   "DB_Inspect_Pistoane_PompaB" : Int = PLC DB_Inspect_Pistoane.Piston_A AT %DB34.DBW28, 1 s
   "DB_Inspect_Pistoane_PompaC" : Int = PLC DB_Inspect_Pistoane.Piston_B AT %DB34.DBW30, 1 s
   "DB_Inspect_Pistoane_CutP1" : Bool = PLC DB_Inspect_Pistoane.Piston_C AT %DB34.DBX32.5, 1 s
   "DB_Inspect_Pistoane_StatusPump1" : Int = PLC DB_Inspect_Pistoane.Presiune_1 AT %DB34.DBW34, 1 s
   "DB_Vizibilitati_Platforme/Colete_Platforma_Rebut" : Bool = PLC DB_Inspect_Pistoane.Presiune_2 AT %DB1.DBX1.0, 100 ms
   "DB_Vizibilitati_Platforme/Colete_Colet_Rebut" : Bool = PLC DB_Inspect_Pistoane.Presiune_A AT %DB1.DBX0.7, 100 ms
   "DB_Tip_Cutie_BoxStatus" : Bool = PLC DB_Inspect_Pistoane.Presiune_B AT %DB37.DBX6.3, 100 ms
   "DB_ControlEnable_ControlEnable_Btn_A" : Bool = PLC DB_Inspect_Pistoane.Presiune_C AT %DB45.DBX0.0, 1 s
   "DB_ControlEnable_ControlEnable_Btn_B" : Bool = PLC DB_Inspect_Pistoane.Presiune_Upper_2 AT %DB45.DBX0.1, 1 s
   "DB_ControlEnable_ControlEnable_Btn_C" : Bool = PLC DB_Inspect_Pistoane.Presiune_Upper_1 AT %DB45.DBX0.2, 1 s
   "DB_ControlEnable_ControlEnable_Btn_Load" : Bool = PLC DB_Inspect_Pistoane.Presiune_Lower_1 AT %DB45.DBX0.3, 1 s
   "DB_ControlEnable_ControlEnable_Btn_ACKLoad" : Bool = PLC DB_Inspect_Pistoane.Presiune_Lower_2 AT %DB45.DBX0.4, 1 s
   "DB_ControlEnable_ControlEnable_Btn_PlaceBox" : Bool = PLC DB_Status_Motoare.Motor_1 AT %DB45.DBX0.6, 1 s
   "DB_general_Piston_Scrap" : Int = PLC DB_HMI.Viz_Platforma_Libera AT %DB2.DBW36, 100 ms
   "DB_Tranzitii_Viz_CutieScrapP3" : Bool = PLC DB_general.Piston_Incarcare AT %DB47.DBX8.0, 100 ms
   "DB_Banda3_AckScrap" : Bool = PLC DB_Banda3.AckScrap AT %DB49.DBX2.1, 100 ms
   "DB_Banda3_Poz_Banda3" : Int = PLC DB_Banda3.Poz_Banda3 AT %DB49.DBW0, 100 ms
   "DB_Banda3_Viz_CutieBanda3" : Bool = PLC DB_Banda3.Viz_CutieBanda3 AT %DB49.DBX2.0, 100 ms
   "DB_HMI_Eng/Ger" : Bool = PLC DB_HMI.Eng AT %DB19.DBX124.0, 1 s
   "DB_HMI_Ger" : Bool = PLC DB_HMI.Ger AT %DB19.DBX138.0, 1 s
   "DB_RemoteAcces_ControlEnable_Stop" : Bool = PLC DB_RemoteAcces.ControlEnable_Stop AT %DB6.DBX0.6, 1 s
   "DB_RemoteAcces_ControlEnable_Start" : Bool = PLC DB_RemoteAcces.ControlEnable_Start AT %DB6.DBX0.7, 1 s
   "DB_RemoteAcces_ControlEnable_Man/Auto" : Bool = PLC DB_RemoteAcces.ControlEnable_Man/Auto AT %DB6.DBX1.0, 1 s
   "DB_ControlEnable_ControlEnable_StartSim" : Bool = PLC DB_ControlEnable.ControlEnable_StartSim AT %DB45.DBX0.5, 1 s
   "DB_SIM_Ack_Load_Pressed" : Bool = PLC DB_SIM.Ack_Load_Pressed AT %DB40.DBX0.3, 1 s
   "DB_ControlEnable_StatusLoadBtn" : Int = PLC DB_ControlEnable.StatusLoadBtn AT %DB45.DBW2, 1 s

HMI tags "Vizibilitate_Log"
   "Viz_Pachet_1" : Bool, internal
   "Viz_Pachet_2" : Bool, internal
   "Viz_Pachet_3" : Bool, internal
   "Viz_Pachet_4" : Bool, internal
   "Viz_Pachet_5" : Bool, internal
   "Viz_Pachet_6" : Bool, internal
   "Viz_Pachet_7" : Bool, internal
   "Viz_Pachet_8" : Bool, internal
   "Viz_Pachet_9" : Bool, internal
   "Viz_Pachet_10" : Bool, internal
   "QR_En" : Bool, internal

HMI tags "DB_HMI_tags"
   "DB_HMI_A_Pressed" : Bool = PLC DB_HMI.A_Pressed AT %DB19.DBX6.0, 100 ms
   "DB_HMI_Ack_Load" : Bool = PLC DB_HMI.Ack_Load AT %DB19.DBX14.3, 100 ms
   "DB_HMI_Add_Ulei" : Bool = PLC DB_HMI.Add_Ulei AT %DB19.DBX42.0, 100 ms
   "DB_HMI_B_Pressed" : Bool = PLC DB_HMI.B_Pressed AT %DB19.DBX6.1, 100 ms
   "DB_HMI_C_Pressed" : Bool = PLC DB_HMI.C_Pressed AT %DB19.DBX6.2, 100 ms
   "DB_HMI_Cutie_Automata" : Bool = PLC DB_HMI.Cutie_Automata AT %DB19.DBX6.3, 100 ms
   "DB_HMI_Cutie_Manuala" : Bool = PLC DB_HMI.Cutie_Manuala AT %DB19.DBX6.4, 100 ms
   "DB_HMI_Greutate" : Real = PLC DB_HMI.Greutate AT %DB19.DBD54, 100 ms
   "DB_HMI_LOAD" : Int = PLC DB_HMI.LOAD AT %DB19.DBW12, 100 ms
   "DB_HMI_LOAD_A" : Bool = PLC DB_HMI.LOAD_A AT %DB19.DBX28.0, 100 ms
   "DB_HMI_LOAD_B" : Bool = PLC DB_HMI.LOAD_B AT %DB19.DBX28.1, 100 ms
   "DB_HMI_LOAD_C" : Bool = PLC DB_HMI.LOAD_C AT %DB19.DBX28.2, 100 ms
   "DB_HMI_Load_RDY" : Bool = PLC DB_HMI.Load_RDY AT %DB19.DBX20.0, 100 ms
   "DB_HMI_Piston_1_Status" : Int = PLC DB_HMI.Piston_1_Status AT %DB19.DBW16, 100 ms
   "DB_HMI_Piston_2_Status" : Int = PLC DB_HMI.Piston_2_Status AT %DB19.DBW18, 100 ms
   "DB_HMI_Racire_Ulei" : Bool = PLC DB_HMI.Racire_Ulei AT %DB19.DBX42.3, 100 ms
   "DB_HMI_Sageata_Deplasare_Banda_Bile" : Bool = PLC DB_HMI.Sageata_Deplasare_Banda_Bile AT %DB19.DBX32.0, 100 ms
   "DB_HMI_Set_T0" : Bool = PLC DB_HMI.Set_T0 AT %DB19.DBX42.6, 100 ms
   "DB_HMI_Set_T50" : Bool = PLC DB_HMI.Set_T50 AT %DB19.DBX42.7, 100 ms
   "DB_HMI_START_SIM" : Bool = PLC DB_HMI.START_SIM AT %DB19.DBX43.0, 100 ms
   "DB_HMI_Start_System" : Bool = PLC DB_HMI.Start_System AT %DB19.DBX42.2, 100 ms
   "DB_HMI_Status_Banda_Bile" : Int = PLC DB_HMI.Status_Banda_Bile AT %DB19.DBW30, 100 ms
   "DB_HMI_Status_Incalzire/Racire_Ulei" : Int = PLC DB_HMI.Status_Incalzire/Racire_Ulei AT %DB19.DBW44, 100 ms
   "DB_HMI_Status_Piston_A" : Int = PLC DB_HMI.Status_Piston_A AT %DB19.DBW22, 100 ms
   "DB_HMI_Status_Piston_B" : Int = PLC DB_HMI.Status_Piston_B AT %DB19.DBW24, 100 ms
   "DB_HMI_Status_Piston_C" : Int = PLC DB_HMI.Status_Piston_C AT %DB19.DBW26, 100 ms
   "DB_HMI_Sub_Ulei" : Bool = PLC DB_HMI.Sub_Ulei AT %DB19.DBX42.1, 100 ms
   "DB_HMI_Temp_Ulei" : Int = PLC DB_HMI.Temp_Ulei AT %DB19.DBW34, 100 ms
   "DB_HMI_TEST_LOAD" : Bool = PLC DB_HMI.BTN_LOAD AT %DB19.DBX43.1, 100 ms
   "DB_HMI_Tip_Cutie" : Int = PLC DB_HMI.Tip_Cutie_Lung AT %DB19.DBW8, 100 ms
   "DB_HMI_Tip_Cutie_Scurt" : Int = PLC DB_HMI.Tip_Cutie_Scurt AT %DB19.DBW10, 100 ms
   "DB_HMI_Transport" : Bool = PLC DB_HMI.Transport AT %DB19.DBX14.0, 100 ms
   "DB_HMI_Ventilator_Cald" : Int = PLC DB_HMI.Ventilator_Cald AT %DB19.DBW50, 100 ms
   "DB_HMI_Ventilator_Rece" : Int = PLC DB_HMI.Ventilator_Rece AT %DB19.DBW48, 100 ms
   "DB_HMI_Viz_Cutie_A" : Bool = PLC DB_HMI.Viz_Cutie_A AT %DB19.DBX20.1, 100 ms
   "DB_HMI_Viz_Cutie_B" : Bool = PLC DB_HMI.Viz_Cutie_B AT %DB19.DBX20.2, 100 ms
   "DB_HMI_Viz_Cutie_Banda_1" : Bool = PLC DB_HMI.Viz_Cutie_Banda_1 AT %DB19.DBX14.2, 100 ms
   "DB_HMI_Viz_Cutie_C" : Bool = PLC DB_HMI.Viz_Cutie_C AT %DB19.DBX20.3, 100 ms
   "DB_HMI_Viz_Cutie_Lunga" : Bool = PLC DB_HMI.Viz_Cutie_Lunga AT %DB19.DBX6.6, 100 ms
   "DB_HMI_Viz_Cutie_Man/Auto" : Int = PLC DB_HMI.Viz_Cutie_Man/Auto AT %DB19.DBW46, 100 ms
   "DB_HMI_Viz_Cutie_Scurta" : Bool = PLC DB_HMI.Viz_Cutie_Scurta AT %DB19.DBX6.5, 100 ms
   "DB_HMI_Viz_Platforma_Libera" : Bool = PLC DB_HMI.Viz_Platforma_Libera AT %DB19.DBX52.0, 100 ms
   "DB_HMI_Volum_Ulei" : Int = PLC DB_HMI.Volum_Ulei AT %DB19.DBW40, 1 s

HMI tags "Alarme"
   "DB_Alarme_Emg_Stop" : Int = PLC DB_Alarme.Emg_Stop AT %DB46.DBW0, Cycle_1

HMI tags "DB_General_tags"
   "DB_general_Piston_2_Cursa_Completa" : Int = PLC DB_general.Piston_2_Cursa_Completa AT %DB2.DBW18, Cycle_1
   "DB_general_Piston_Cursa_Completa" : Int = PLC DB_general.Piston_1_Cursa_Completa AT %DB2.DBW16, 100 ms
   "DB_general_Piston_Incarcare" : Int = PLC DB_general.Piston_Incarcare AT %DB2.DBW28, 100 ms
   "DB_general_Piston_Incarcare_A" : Int = PLC DB_general.Piston_Incarcare_A AT %DB2.DBW30, 100 ms
   "DB_general_Piston_Incarcare_B" : Int = PLC DB_general.Piston_Incarcare_B AT %DB2.DBW32, 100 ms
   "DB_general_Piston_Incarcare_C" : Int = PLC DB_general.Piston_Incarcare_C AT %DB2.DBW34, 100 ms
   "DB_general_Poz_Cutie_Bile" : Int = PLC DB_general.Poz_Cutie_Bile AT %DB2.DBW8, 100 ms
   "DB_general_Poz_Piston_1" : Int = PLC DB_general.Poz_Piston_1 AT %DB2.DBW2, 100 ms
   "DB_general_Senzor_1_Descarcare" : Bool = PLC DB_general.Senzor_1_Descarcare AT %DB2.DBX0.4, 100 ms
   "DB_general_Senzor_1_Incarcare" : Bool = PLC DB_general.Senzor_1_Incarcare AT %DB2.DBX0.2, 100 ms
   "DB_general_Senzor_2_Incarcare" : Bool = PLC DB_general.Senzor_2_Incarcare AT %DB2.DBX0.3, 100 ms
   "DB_general_Stare_Poz_Incarcare" : Bool = PLC DB_general.Stare_Poz_Incarcare AT %DB2.DBX0.0, 100 ms
   "DB_general_Valoare" : Int = PLC DB_general.Valoare AT %DB2.DBW14, 100 ms

HMI tags "DB_Inspect_tags"
   "DB_Inspect_Pistoane_Piston_1" : Bool = PLC DB_Inspect_Pistoane.Piston_1 AT %DB34.DBX0.0, 1 s
   "DB_Inspect_Pistoane_Piston_2" : Bool = PLC DB_Inspect_Pistoane.Piston_2 AT %DB34.DBX0.1, 1 s
   "DB_Inspect_Pistoane_Piston_A" : Bool = PLC DB_Inspect_Pistoane.Piston_A AT %DB34.DBX0.2, 1 s
   "DB_Inspect_Pistoane_Piston_B" : Bool = PLC DB_Inspect_Pistoane.Piston_B AT %DB34.DBX0.3, 1 s
   "DB_Inspect_Pistoane_Piston_C" : Bool = PLC DB_Inspect_Pistoane.Piston_C AT %DB34.DBX0.4, 1 s
   "DB_Inspect_Pistoane_Presiune_1" : Int = PLC DB_Inspect_Pistoane.Presiune_1 AT %DB34.DBW2, 1 s
   "DB_Inspect_Pistoane_Presiune_2" : Int = PLC DB_Inspect_Pistoane.Presiune_2 AT %DB34.DBW4, 1 s
   "DB_Inspect_Pistoane_Presiune_A" : Int = PLC DB_Inspect_Pistoane.Presiune_A AT %DB34.DBW6, 1 s
   "DB_Inspect_Pistoane_Presiune_B" : Int = PLC DB_Inspect_Pistoane.Presiune_B AT %DB34.DBW8, 1 s
   "DB_Inspect_Pistoane_Presiune_C" : Int = PLC DB_Inspect_Pistoane.Presiune_C AT %DB34.DBW10, 1 s
   "DB_Inspect_Pistoane_Presiune_Lower_1" : Int = PLC DB_Inspect_Pistoane.Presiune_Lower_1 AT %DB34.DBW16, 1 s
   "DB_Inspect_Pistoane_Presiune_Lower_2" : Int = PLC DB_Inspect_Pistoane.Presiune_Lower_2 AT %DB34.DBW18, 1 s
   "DB_Inspect_Pistoane_Presiune_Upper_1" : Int = PLC DB_Inspect_Pistoane.Presiune_Upper_1 AT %DB34.DBW14, 1 s
   "DB_Inspect_Pistoane_Presiune_Upper_2" : Int = PLC DB_Inspect_Pistoane.Presiune_Upper_2 AT %DB34.DBW12, 1 s

HMI tags "DB_Status_tags"
   "DB_Status_Motoare_Motor_1" : Int = PLC DB_Status_Motoare.Motor_1 AT %DB25.DBW0, 100 ms
   "DB_Status_Pistoane_Status_Pison_2" : Int = PLC DB_Status_Pistoane.Status_Pison_2 AT %DB26.DBW2, 100 ms
   "DB_Status_Pistoane_Status_Piston_1" : Int = PLC DB_Status_Pistoane.Status_Piston_1 AT %DB26.DBW0, 100 ms
   "DB_Status_Pistoane_Status_Piston_A" : Int = PLC DB_Status_Pistoane.Status_Piston_A AT %DB26.DBW4, 100 ms
   "DB_Status_Pistoane_Status_Piston_B" : Int = PLC DB_Status_Pistoane.Status_Piston_B AT %DB26.DBW6, 100 ms
   "DB_Status_Pistoane_Status_Piston_C" : Int = PLC DB_Status_Pistoane.Status_Piston_C AT %DB26.DBW8, 100 ms

discrete alarms
   1: 'Emergency Stop / Not-Halt', class Errors, trigger "DB_Alarme_Emg_Stop" bit 0
   2: 'The weight tolerance is too high and the intervals overlap / Die Gewichtstoleranz ist zu hoch und die Intervalle überschneiden sich', class Errors, trigger "DB_Tip_Cutie_IntersectieInterval" bit 1
   3: 'The placed box will be cosidered scrap / Die platzierte Kiste gilt als Schrott', class Acknowledgement, trigger "DB_Tip_Cutie_Scrap" bit 0

analog alarms
   8: 'Hydraulic oil volume too low / Hydraulikölmenge zu gering', class Errors, trigger "DB_HMI_Volum_Ulei"
   7: 'Hydraulic oil volume too high / Hydraulikölmenge zu hoch', class Errors, trigger "DB_HMI_Volum_Ulei"
   3: 'No more free spaces in B slot / Keine freien Plätze mehr im B-Steckplatz', class Acknowledgement, trigger "Locuri_B"
   6: 'Hydraulic oil too cold / Hydrauliköl zu kalt', class Errors, trigger "DB_HMI_Temp_Ulei"
   5: 'Hydraulic oil overheated / Hydrauliköl überhitzt', class Errors, trigger "DB_HMI_Temp_Ulei"
   2: 'No more free spaces in A slot / Keine freien Plätze mehr im A-Steckplatz', class Acknowledgement, trigger "Locuri_A"
   4: 'No more free spaces in C slot / Keine freien Plätze mehr im C-Steckplatz / Nu exista locuri disponibile in C / Keine freien Plätze mehr im C-Steckplatz', class Acknowledgement, trigger "Locuri_C"
   1: 'The weight limit on A truck has not been set / Die Gewichtsbeschränkung für A LKW wurde nicht festgelegt', class Errors, trigger "DB_HMI_MaxLoad_A"
   9: 'The weight limit on B truck has not been set / Die Gewichtsbeschränkung für B LKW wurde nicht festgelegt', class Errors, trigger "DB_HMI_MaxLoad_A"
   10: 'The weight limit on C truck has not been set / Die Gewichtsbeschränkung für C LKW wurde nicht festgelegt', class Errors, trigger "DB_HMI_MaxLoad_A"
   11: 'The weight tolerance is too high and the intervals overlap / Die Gewichtstoleranz ist zu hoch und die Intervalle überschneiden sich', class Errors, trigger "DB_general_GreutateMaxManual"
   12: 'The pump 1 is in error state', class Errors, trigger "DB_Inspect_Pistoane_StatusPump1"
   13: 'Unload the box from the conveyor band 3', class Acknowledgement, trigger "DB_Banda3_Poz_Banda3"

graphic list "@DiagnosticsStates": 0 '@Diagnostics_StateGood'; 1 '@Diagnostics_StateBad'

screen "Statie Distribuire" 1920x1080, template "Template_1"
   Visibility <- "DB_Status_Pistoane_Status_Piston_1"
   GraphicView "Graphic view_5" at 1452,223 size 335x213; Picture "background.xwr"
   Rectangle "Rectangle_17" at 1638,184 size 45x71
      VerticalMovement <- "DB_general_Piston_2_Cursa_Completa"
   Rectangle "Rectangle_18" at 1623,184 size 75x71
      VerticalMovement <- "DB_general_Piston_2_Cursa_Completa"
   Rectangle "Rectangle_19" at 1608,184 size 105x71
      VerticalMovement <- "DB_general_Piston_2_Cursa_Completa"
   GraphicView "Graphic view_7" at 770,388 size 329x228; Picture "background.xwr"
   Switch "Switch_6" at 17,754 size 224x133; TextOn 'Placed Box Kolben Status'; CaptionText 'Switch'; TextOff 'Place Box Kolben Status'
      on SwitchOff: SetTag("DB_general_Senzor_1_Incarcare", 0); SetTag("DB_general_Senzor_2_Incarcare", 0)
      on SwitchOn: SetTag("DB_general_Senzor_1_Incarcare", 1); SetTag("DB_general_Senzor_2_Incarcare", 1); SetTag("DB_Tip_Cutie_BoxStatus", 1)
      Appearance <- "DB_HMI_Viz_Cutie_Scurta"
      ProcessValue <- "DB_HMI_Viz_Cutie_Scurta"
      ObjectEnable <- "DB_ControlEnable_ControlEnable_Btn_PlaceBox"
   Switch "Switch_7" at 246,754 size 224x133; TextOn 'ACK LOAD ACK LAST'; CaptionText 'Switch'; TextOff 'ACK LOAD ACK LAST'
      on SwitchOn: SetTag("DB_HMI_Load_RDY", 1)
      ProcessValue <- "DB_HMI_Ack_Load"
      Appearance <- "DB_general_Stare_Poz_Incarcare"
      ObjectEnable <- "DB_ControlEnable_ControlEnable_Btn_ACKLoad"
   Switch "Switch_9" at 477,754 size 269x133; TextOn 'LOAD / BELASTUNG'; CaptionText 'Switch'; TextOff 'LOAD / BELASTUNG'
      ObjectEnable <- "DB_ControlEnable_ControlEnable_Btn_Load"
      ProcessValue <- "DB_HMI_TEST_LOAD"
      Appearance <- "DB_ControlEnable_StatusLoadBtn"
      on SwitchOn: SetTag("DB_ControlEnable_StatusLoadBtn", 1)
      on SwitchOff: SetTag("DB_ControlEnable_StatusLoadBtn", 0)
   Rectangle "Rectangle_8" at 910,550 size 65x71
      VerticalMovement <- "DB_general_Piston_Cursa_Completa"
   Rectangle "Rectangle_7" at 900,550 size 85x71
      VerticalMovement <- "DB_general_Piston_Cursa_Completa"
   Rectangle "Rectangle_6" at 890,550 size 105x71
      VerticalMovement <- "DB_general_Piston_Cursa_Completa"
   Rectangle "Rectangle_10" at 850,530 size 185x25
      VerticalMovement <- "DB_general_Piston_Cursa_Completa"
   TextField "Text field_8" at 1114,477 size 100x50; Text 'S1'
   TextField "Text field_9" at 1111,527 size 100x50; Text 'S2'
   Rectangle "Rectangle_14" at 1044,488 size 45x33
      Appearance <- "DB_general_Senzor_1_Incarcare"
   Rectangle "Rectangle_15" at 1044,536 size 45x33
      Appearance <- "DB_general_Senzor_2_Incarcare"
   Rectangle "Rectangle_16" at 1752,276 size 45x33
      Appearance <- "DB_general_Senzor_1_Descarcare"
   Rectangle "Rectangle_20" at 1752,327 size 45x33
      Appearance <- "DB_general_Senzor_1_Descarcare"
   TextField "Text field_13" at 1807,323 size 76x38; Text 'S4'
   Rectangle "Rectangle_22" at 1568,251 size 175x21
      VerticalMovement <- "DB_general_Piston_2_Cursa_Completa"
   TextField "Text field_5" at 1805,276 size 76x38; Text 'S3'
   Rectangle "Rectangle_24" at 796,626 size 40x37
      Appearance <- "DB_Status_Pistoane_Status_Piston_1"
   TextField "Text field_4" at 802,630 size 52x26; Text 'P1'
   Button "Button_1" at 1182,469 size 371x100; TextOff 'RESET / ZURÜCKSETZEN'
      on Release: SetTag("DB_SIM_BTN_RESET", 0)
      on Press: SetTag("DB_HMI_Viz_Cutie_Scurta", 0); SetTag("LOAD", 0); SetTag("DB_HMI_Ack_Load", 0); SetTag("DB_SIM_BTN_RESET", 1); SetTag("DB_general_Senzor_1_Incarcare", 0); SetTag("DB_general_Senzor_2_Incarcare", 0); SetTag("LOAD", 0); SetTag("DB_HMI_TEST_LOAD", 0); SetTag("DB_HMI_Viz_Cutie_Man/Auto", 0); SetTag("DB_HMI_Viz_Cutie_Banda_1", 0); SetTag("DB_HMI_Greutate", 0); SetTag("DB_HMI_START_SIM", 0); SetTag("DB_HMI_A_Pressed", 0); SetTag("DB_HMI_B_Pressed", 0); SetTag("DB_HMI_C_Pressed", 0); SetTag("DB_SIM_Ack_Load_Pressed", 0)
   GraphicView "Graphic view_6" at 1299,125 size 196x98; Picture "Graphic_76"
   GraphicView "Graphic view_3" at 879,124 size 196x98; Picture "Graphic_76"
   Switch "Switch_1" at 313,462 size 74x60; TextOn 'A'; CaptionText 'Switch'; TextOff 'A'
      on SwitchOff: SetTag("DB_HMI_Viz_Cutie_A", 0)
      on SwitchOn: SetTag("DB_HMI_B_Pressed", 0); SetTag("DB_HMI_C_Pressed", 0); SetTag("DB_HMI_Viz_Cutie_A", 1); SetTag("DB_HMI_Viz_Cutie_B", 0); SetTag("DB_HMI_Viz_Cutie_C", 0)
      Appearance <- "DB_HMI_A_Pressed"
      ProcessValue <- "DB_HMI_A_Pressed"
      ObjectEnable <- "DB_ControlEnable_ControlEnable_Btn_A"
   Switch "Switch_3" at 415,460 size 74x60; TextOn 'B'; CaptionText 'Switch'; TextOff 'B'
      on SwitchOn: SetTag("DB_HMI_A_Pressed", 0); SetTag("DB_HMI_C_Pressed", 0); SetTag("DB_HMI_Viz_Cutie_B", 1); SetTag("DB_HMI_Viz_Cutie_A", 0); SetTag("DB_HMI_Viz_Cutie_C", 0)
      Appearance <- "DB_HMI_B_Pressed"
      ProcessValue <- "DB_HMI_B_Pressed"
      ObjectEnable <- "DB_ControlEnable_ControlEnable_Btn_B"
   Switch "Switch_4" at 524,460 size 74x60; TextOn 'C'; CaptionText 'Switch'; TextOff 'C'
      on SwitchOn: SetTag("DB_HMI_A_Pressed", 0); SetTag("DB_HMI_B_Pressed", 0); SetTag("DB_HMI_Viz_Cutie_C", 1); SetTag("DB_HMI_Viz_Cutie_B", 0); SetTag("DB_HMI_Viz_Cutie_A", 0)
      Appearance <- "DB_HMI_C_Pressed"
      ProcessValue <- "DB_HMI_C_Pressed"
      ObjectEnable <- "DB_ControlEnable_ControlEnable_Btn_C"
   TextField "Text field_17" at 125,420 size 185x40; Text 'Weight / Gewicht'
   TextField "Text field_3" at 354,417 size 255x34; Text 'Destination / Ziel'
   IOField "I/O field_2" at 310,526 size 46x49; FormatPattern 9
      ProcessValue <- "Locuri_A"
   IOField "I/O field_3" at 425,526 size 46x49; FormatPattern 9
      ProcessValue <- "Locuri_B"
   IOField "I/O field_4" at 535,529 size 46x49; FormatPattern 9
      ProcessValue <- "Locuri_C"
   IOField "I/O field_1" at 115,491 size 144x59; FormatPattern 999; Unit  Kg
      ProcessValue <- "DB_HMI_Greutate"
   Rectangle "Rectangle_30" at 1619,138 size 40x37
      Appearance <- "DB_Status_Pistoane_Status_Pison_2"
   TextField "Text field_6" at 1625,142 size 46x26; Text 'P2'
   Rectangle "Rectangle_26" at 962,171 size 53x44
      Appearance <- "DB_Status_Motoare_Motor_1"
   Rectangle "Rectangle_29" at 1380,171 size 53x44
      Appearance <- "DB_Status_Motoare_Motor_1"
   Switch "Switch_8" at 1138,592 size 345x100; CaptionText 'Switch'; TextOff 'Start Sim / Starten Sie Sim'; TextOn 'Started Sim / Sim gestartet'
      Visibility <- "Man/Auto"
      ProcessValue <- "DB_HMI_START_SIM"
   TextField "Text field_10" at 968,172 size 82x32; Text 'M1'
   TextField "Text field_11" at 1383,175 size 82x32; Text 'M2'
   GraphicView "Graphic view_4" at 870,410 size 145x119; Picture "Box"
      Visibility <- "DB_Tranzitii_Viz_Cutie_1"
      VerticalMovement <- "DB_general_Piston_Cursa_Completa"
   GraphicView "Graphic view_1" at 1582,280 size 145x119; Picture "Box"
      Visibility <- "DB_Tranzitii_VizCutieEnd"
      VerticalMovement <- "DB_general_Piston_2_Cursa_Completa"
   TextField "Text field_21" at 88,80 size 608x40; Text 'REMOTE EMG/STOP/START / FERN-EMG/STOP/START'
   Switch "Switch_2" at 97,148 size 150x76; CaptionText 'Switch'; TextOff 'EMG'; TextOn 'EMG'
      ProcessValue <- "DB_RemoteAcces_EmgStopBtn"
      Appearance <- "DB_RemoteAcces_EmgStopBtn"
      on SwitchOn: SetTag("DB_RemoteAcces_On/Off", 0)
   Button "Button_3" at 274,148 size 152x77; TextOff 'Stop'
      on Click: SetTag("DB_RemoteAcces_On/Off", 0)
      Appearance <- "DB_RemoteAcces_On/Off"
      ObjectEnable <- "DB_RemoteAcces_ControlEnable_Stop"
   Button "Button_4" at 447,149 size 155x76; TextOff 'Start'
      on Click: SetTag("DB_RemoteAcces_On/Off", 1)
      Appearance <- "DB_RemoteAcces_On/Off"
      ObjectEnable <- "DB_RemoteAcces_ControlEnable_Start"
   Switch "Switch_5" at 101,243 size 255x53; CaptionText 'Switch'; TextOff 'Automat / Automatisch'; TextOn 'Manual / manuell'
      ProcessValue <- "DB_RemoteAcces_Manual/Auto"
      ObjectEnable <- "DB_RemoteAcces_ControlEnable_Man/Auto"
   Switch "Switch_10" at 369,246 size 233x53; CaptionText 'Switch'; TextOff 'Local / Lokal'; TextOn 'Remote / Fern'; Authorization "Monitor"
      ProcessValue <- "DB_RemoteAcces_Remote"
   Switch "Switch_11" at 1502,592 size 372x100; TextOn 'Started Sim / Sim gestartet'; CaptionText 'Switch'; TextOff 'Start Sim / Starten Sie Sim'
      ProcessValue <- "DB_HMI_START_SIM"
      Visibility <- "DB_RemoteAcces_Manual/Auto"
      ObjectEnable <- "DB_ControlEnable_ControlEnable_StartSim"
   GraphicView "Graphic view_2" at 870,276 size 145x119; Picture "Box"
      HorizontalMovement <- "Poz_Cutie"
      Visibility <- "DB_HMI_Viz_Cutie_Banda_1"
   Switch "Switch_16" at 775,730 size 364x53; TextOn 'Box in transit / Box im Transport'; CaptionText 'Switch'; TextOff 'Waiting for box / Warten auf die Kiste'
      ProcessValue <- "DB_Tip_Cutie_BoxStatus"
   Switch "Switch_17" at 1151,730 size 178x53; TextOn 'Weight / Gewicht'; CaptionText 'Switch'; TextOff 'Weight / Gewicht'
   Switch "Switch_18" at 1341,730 size 357x53; TextOn 'Type of gearbox / Getriebetyp'; CaptionText 'Switch'; TextOff 'Type of gearbox / Getriebetyp'
   Switch "Switch_19" at 1382,788 size 255x42; TextOn 'Manual / manuell'; CaptionText 'Switch'; TextOff 'Automatic / Automatikgetriebe'
      ProcessValue <- "DB_Tip_Cutie_TipCutie"
      Visibility <- "DB_Tip_Cutie_VizTipCutie"
   Switch "Switch_12" at 1351,788 size 337x42; TextOn 'Scrap / Schrott'; CaptionText 'Switch'; TextOff 'Scrap / Schrott'
      ProcessValue <- "DB_Tip_Cutie_TipCutie"
      Visibility <- "DB_Tip_Cutie_RebutLbl"
   IOField "I/O field_5" at 1173,788 size 151x45; Authorization "Monitor"; FormatPattern 999; Unit  Kg
      ProcessValue <- "DB_HMI_Greutate"

Template "Template_1" 1920x1080
   Button "Template_Button_4" at 1158,932 size 290x140; TextOff 'Packets Log Pakete Protokoll'
      on Click: ActivateScreen("Log_Cutii", 0); SetTag("Template_Satie_Distribuire", 0); SetTag("Template_Statie_Incarcare", 0); SetTag("Template_Packets_Log", 1); SetTag("Template_Hidraulic_Station", 0); SetTag("Template_Errors", 0); SetTag("Template_Home", 0)
      Appearance <- "Template_Packets_Log"
   Button "Template_Button_7" at 556,930 size 293x140; TextOff 'Loading Station Lade- station'
      on Click: ActivateScreen("Statie Incarcare", 0); SetTag("Template_Satie_Distribuire", 0); SetTag("Template_Statie_Incarcare", 1); SetTag("Template_Packets_Log", 0); SetTag("Template_Hidraulic_Station", 0); SetTag("Template_Errors", 0); SetTag("Template_Home", 0)
      Appearance <- "Template_Statie_Incarcare"
   Button "Template_Button_8" at 857,931 size 295x140; TextOff 'Hydraulic Station Hydraulik- station'
      on Click: ActivateScreen("Statie Hidraulica", 0); SetTag("Template_Satie_Distribuire", 0); SetTag("Template_Statie_Incarcare", 0); SetTag("Template_Packets_Log", 0); SetTag("Template_Hidraulic_Station", 1); SetTag("Template_Errors", 0); SetTag("Template_Home", 0)
      Appearance <- "Template_Hidraulic_Station"
   Button "Template_Button_9" at 224,930 size 323x140; TextOff 'Distribution Station Verteiler- station'
      on Click: ActivateScreen("Statie Distribuire", 0); SetTag("Template_Satie_Distribuire", 1); SetTag("Template_Statie_Incarcare", 0); SetTag("Template_Packets_Log", 0); SetTag("Template_Hidraulic_Station", 0); SetTag("Template_Errors", 0); SetTag("Template_Home", 0)
      Appearance <- "Template_Satie_Distribuire"
   Button "Template_Button_10" at 1458,931 size 142x138; TextOff 'Back / Zurück'
      on Click: function_efd93a16()
   Button "Template_Button_5" at 1609,934 size 142x135; TextOff 'Text'
      on Click: ActivateScreen("Alarme", 0); SetTag("Template_Home", 0); SetTag("Template_Satie_Distribuire", 0); SetTag("Template_Statie_Incarcare", 0); SetTag("Template_Packets_Log", 0); SetTag("Template_Hidraulic_Station", 0); SetTag("Template_Errors", 1); SetTag("Template_Home", 0)
      Appearance <- "Template_Errors"
   GraphicView "Template_Graphic view_1" at 1634,955 size 86x91; Picture "Graphic_73"
   Button "Template_Button_1" at 5,931 size 203x140; TextOff 'Text'
      on Click: ActivateScreen("Home", 0); SetTag("Template_Satie_Distribuire", 0); SetTag("Template_Statie_Incarcare", 0); SetTag("Template_Packets_Log", 0); SetTag("Template_Hidraulic_Station", 0); SetTag("Template_Errors", 0); SetTag("Template_Home", 1)
      Appearance <- "Template_Home"
   GraphicView "Template_Graphic view_2" at 41,957 size 122x89; Picture "Graphic_112"
   GraphicView "Template_Graphic view_4" at 1718,0 size 202x110; Picture "Color-Siemens-Logo"
   Button "Template_Button_2" at 1760,932 size 142x134; TextOff 'Text'
      on Release: StopRuntime(0)
   GraphicView "Template_Graphic view_3" at 1788,962 size 85x73; Picture "Graphic_113"

screen "Home" 1920x1080, template "Template_1"
   on GenerateScreen: function_f23ef4c9(); SetTag("Template_Satie_Distribuire", 0); SetTag("Template_Statie_Incarcare", 0); SetTag("Template_Packets_Log", 0); SetTag("Template_Hidraulic_Station", 0); SetTag("Template_Errors", 0)
   GraphicView "Graphic view_16" at 566,192 size 257x175; Picture "background.xwr"
   GraphicView "Graphic view_18" at 557,745 size 257x175; Picture "background.xwr"
   GraphicView "Graphic view_5" at 572,81 size 257x175; Picture "background.xwr"
   Rectangle "Rectangle_51" at 674,251 size 107x95
      VerticalMovement <- "DB_general_Poz_Cutie_Bile"
      Visibility <- "DB_Vizibilitati_Platforme/Colete_Platforma_Rebut"
   Rectangle "Rectangle_64" at 841,851 size 57x22
      HorizontalMovement <- "DB_general_Piston_Scrap"
   Rectangle "Rectangle_78" at 841,849 size 57x26
      HorizontalMovement <- "DB_general_Piston_Scrap"
   Rectangle "Rectangle_79" at 841,844 size 57x36
      HorizontalMovement <- "DB_general_Piston_Scrap"
   Rectangle "Rectangle_80" at 842,837 size 57x49
      HorizontalMovement <- "DB_general_Piston_Scrap"
   Switch "Switch_1" at 107,707 size 203x48; TextOn 'ACK SCRAP / ACK DEFEKT'; CaptionText 'Switch'; TextOff 'ACK SCRAP / ACK DEFEKT'
      ProcessValue <- "DB_Banda3_AckScrap"
      Appearance <- "DB_Banda3_AckScrap"
   Rectangle "Rectangle_23" at 674,251 size 107x95
      VerticalMovement <- "DB_general_Poz_Cutie_Bile"
      Visibility <- "DB_Vizibilitati_Platforme/Colete_Platforma_C"
   Rectangle "Rectangle_25" at 674,251 size 107x95
      VerticalMovement <- "DB_general_Poz_Cutie_Bile"
      Visibility <- "DB_Vizibilitati_Platforme/Colete_Platforma_B"
   Rectangle "Rectangle_48" at 674,251 size 107x95
      Visibility <- "DB_HMI_Viz_Platforma_Libera"
      VerticalMovement <- "DB_general_Poz_Cutie_Bile"
   Rectangle "Rectangle_12" at 674,251 size 107x95
      VerticalMovement <- "DB_general_Poz_Cutie_Bile"
      Visibility <- "DB_Vizibilitati_Platforme/Colete_Platforma_A"
   Rectangle "Rectangle_52" at 720,50 size 21x58
      VerticalMovement <- "DB_general_Piston_2_Cursa_Completa"
   Rectangle "Rectangle_17" at 712,49 size 38x58
      VerticalMovement <- "DB_general_Piston_2_Cursa_Completa"
   Rectangle "Rectangle_18" at 703,49 size 58x58
      VerticalMovement <- "DB_general_Piston_2_Cursa_Completa"
   Rectangle "Rectangle_19" at 691,49 size 81x58
      VerticalMovement <- "DB_general_Piston_2_Cursa_Completa"
   GraphicView "Graphic view_1" at 686,259 size 84x80; Picture "Box"
      VerticalMovement <- "DB_general_Poz_Cutie_Bile"
      Visibility <- "DB_Vizibilitati_Platforme/Colete_Colet_C"
   GraphicView "Graphic view_12" at 686,259 size 84x80; Picture "Box"
      VerticalMovement <- "DB_general_Poz_Cutie_Bile"
      Visibility <- "DB_Vizibilitati_Platforme/Colete_Colet_B"
   GraphicView "Graphic view_13" at 686,259 size 84x80; Picture "Box"
      VerticalMovement <- "DB_general_Poz_Cutie_Bile"
      Visibility <- "DB_Vizibilitati_Platforme/Colete_Colet_A"
   Rectangle "Rectangle_27" at 557,555 size 72x29
      HorizontalMovement <- "DB_general_Piston_Incarcare_B"
   Rectangle "Rectangle_28" at 557,552 size 72x34
      HorizontalMovement <- "DB_general_Piston_Incarcare_B"
   Rectangle "Rectangle_31" at 560,546 size 72x46
      HorizontalMovement <- "DB_general_Piston_Incarcare_B"
   Rectangle "Rectangle_32" at 557,537 size 72x63
      HorizontalMovement <- "DB_general_Piston_Incarcare_B"
   GraphicView "Graphic view_7" at 48,216 size 253x187; Picture "background.xwr"
   GraphicView "Graphic view_4" at 135,253 size 84x80; Picture "Box"
      Visibility <- "DB_Tranzitii_Viz_Cutie_1"
      VerticalMovement <- "DB_general_Piston_Cursa_Completa"
   Rectangle "Rectangle_33" at 557,711 size 72x29
      HorizontalMovement <- "DB_general_Piston_Incarcare_C"
   Rectangle "Rectangle_34" at 557,708 size 72x34
      HorizontalMovement <- "DB_general_Piston_Incarcare_C"
   Rectangle "Rectangle_35" at 560,702 size 72x46
      HorizontalMovement <- "DB_general_Piston_Incarcare_C"
   Rectangle "Rectangle_36" at 557,693 size 72x63
      HorizontalMovement <- "DB_general_Piston_Incarcare_C"
   Rectangle "Rectangle_37" at 557,412 size 72x29
      HorizontalMovement <- "DB_general_Piston_Incarcare_A"
   Rectangle "Rectangle_38" at 557,409 size 72x34
      HorizontalMovement <- "DB_general_Piston_Incarcare_A"
   Rectangle "Rectangle_39" at 560,403 size 72x46
      HorizontalMovement <- "DB_general_Piston_Incarcare_A"
   Rectangle "Rectangle_40" at 557,394 size 72x63
      HorizontalMovement <- "DB_general_Piston_Incarcare_A"
   GraphicView "Graphic view_2" at 135,138 size 84x80; Picture "Box"
      HorizontalMovement <- "Poz_Cutie"
      Visibility <- "DB_HMI_Viz_Cutie_Banda_1"
   Rectangle "Rectangle_8" at 155,349 size 50x58
      VerticalMovement <- "DB_general_Piston_Cursa_Completa"
   Rectangle "Rectangle_7" at 148,349 size 65x58
      VerticalMovement <- "DB_general_Piston_Cursa_Completa"
   Rectangle "Rectangle_6" at 140,349 size 81x58
      VerticalMovement <- "DB_general_Piston_Cursa_Completa"
   Rectangle "Rectangle_10" at 109,338 size 142x16
      VerticalMovement <- "DB_general_Piston_Cursa_Completa"
   TextField "Text field_8" at 312,289 size 76x38; Text 'S1'
   TextField "Text field_9" at 310,330 size 76x38; Text 'S2'
   Rectangle "Rectangle_14" at 258,298 size 30x26
      Appearance <- "DB_general_Senzor_1_Incarcare"
   Rectangle "Rectangle_15" at 258,338 size 30x26
      Appearance <- "DB_general_Senzor_2_Incarcare"
   Rectangle "Rectangle_16" at 802,125 size 30x26
      Appearance <- "DB_general_Senzor_1_Descarcare"
   Rectangle "Rectangle_20" at 802,167 size 30x26
      Appearance <- "DB_general_Senzor_1_Descarcare"
   Rectangle "Rectangle_22" at 661,104 size 134x16
      VerticalMovement <- "DB_general_Piston_2_Cursa_Completa"
   TextField "Text field_5" at 841,116 size 76x38; Text 'S3'
   Rectangle "Rectangle_24" at 68,412 size 31x30
      Appearance <- "DB_Status_Pistoane_Status_Piston_1"
   TextField "Text field_4" at 74,416 size 38x20; Text 'P1'
   GraphicView "Graphic view_6" at 454,1 size 150x80; Picture "Graphic_76"
   GraphicView "Graphic view_3" at 132,0 size 150x80; Picture "Graphic_76"
   Rectangle "Rectangle_30" at 700,11 size 31x30
      Appearance <- "DB_Status_Pistoane_Status_Pison_2"
   TextField "Text field_6" at 706,15 size 34x20; Text 'P2'
   Rectangle "Rectangle_26" at 195,39 size 41x36
      Appearance <- "DB_Status_Motoare_Motor_1"
   Rectangle "Rectangle_29" at 516,39 size 41x36
      Appearance <- "DB_Status_Motoare_Motor_1"
   TextField "Text field_10" at 199,43 size 69x26; Text 'M1'
   TextField "Text field_11" at 520,43 size 69x26; Text 'M2'
   GraphicView "Graphic view_8" at 813,365 size 450x138; Picture "Graphic_30"
   GraphicView "Graphic view_9" at 811,510 size 450x138; Picture "Graphic_30"
   GraphicView "Graphic view_10" at 810,668 size 450x138; Picture "Graphic_30"
   Rectangle "Rectangle_58" at 622,375 size 24x106
      HorizontalMovement <- "DB_general_Piston_Incarcare_A"
   Rectangle "Rectangle_68" at 622,674 size 24x106
      HorizontalMovement <- "DB_general_Piston_Incarcare_C"
   Rectangle "Rectangle_69" at 481,410 size 68x37
      Appearance <- "DB_Status_Pistoane_Status_Piston_A"
   Rectangle "Rectangle_70" at 481,561 size 68x37
      Appearance <- "DB_Status_Pistoane_Status_Piston_B"
   Rectangle "Rectangle_71" at 480,712 size 68x37
      Appearance <- "DB_Status_Pistoane_Status_Piston_C"
   TextField "Text field_1" at 490,712 size 74x32; Text 'P-C'
   TextField "Text field_2" at 490,558 size 81x32; Text 'P-B'
   TextField "Text field_3" at 489,410 size 74x32; Text 'P-A'
   TextField "Text field_13" at 841,161 size 76x38; Text 'S4'
   Button "Button_1" at 1394,387 size 351x76; TextOff 'Log In Admin / Login-Administrator'; Authorization "User administration"
      on Change: ActivateScreen("AdminPage", 0)
      on Click: SetTag("Template_Home", 0); SetTag("Template_Satie_Distribuire", 0); SetTag("Template_Statie_Incarcare", 0); SetTag("Template_Packets_Log", 0); SetTag("Template_Hidraulic_Station", 0); SetTag("Template_Errors", 0)
   GraphicView "Graphic view_17" at 686,138 size 84x80; Picture "Box"
      VerticalMovement <- "DB_general_Piston_2_Cursa_Completa"
      Visibility <- "DB_Tranzitii_VizCutieEnd"
   TextField "Text field_18" at 770,405 size 263x40; Text 'Available places / Verfügbare Plätze'
   IOField "I/O field_1" at 1041,401 size 58x24; FormatPattern 999
      ProcessValue <- "Locuri_A"
   TextField "Text field_19" at 772,547 size 267x40; Text 'Available places / Verfügbare Plätze'
   IOField "I/O field_2" at 1037,547 size 58x24; FormatPattern 999
      ProcessValue <- "Locuri_B"
   TextField "Text field_20" at 778,705 size 275x40; Text 'Available places / Verfügbare Plätze'
   IOField "I/O field_3" at 1037,707 size 58x24; FormatPattern 999
      ProcessValue <- "Locuri_C"
   Rectangle "Rectangle_50" at 622,518 size 24x106
      HorizontalMovement <- "DB_general_Piston_Incarcare_B"
   GraphicView "Graphic view_20" at 3,798 size 114x126; Picture "Graphic_116"
   GraphicView "Graphic view_19" at 686,822 size 84x80; Picture "Box"
      HorizontalMovement <- "DB_general_Piston_Scrap"
      Visibility <- "DB_Tranzitii_Viz_CutieScrapP3"
   GraphicView "Graphic view_21" at 576,822 size 84x80; Picture "Box"
      HorizontalMovement <- "DB_Banda3_Poz_Banda3"
      Visibility <- "DB_Banda3_Viz_CutieBanda3"
   GraphicView "Graphic view_11" at 686,259 size 84x80; Picture "Box"
      VerticalMovement <- "DB_general_Poz_Cutie_Bile"
      Visibility <- "DB_Vizibilitati_Platforme/Colete_Colet_Rebut"
   Rectangle "Rectangle_82" at 826,821 size 19x82
      HorizontalMovement <- "DB_general_Piston_Scrap"
   Button "Button_2" at 97,705 size 225x51; TextOff 'ACK SCRAP / ACK DEFEKT'
      on Press: SetTag("DB_Banda3_AckScrap", 1)
      on Release: SetTag("DB_Banda3_AckScrap", 0)
   GraphicView "Graphic view_23" at 1688,518 size 159x88; Picture "Graphic_125"
   Button "Button_6" at 1687,518 size 160x88; TextOff 'Text'
      on Click: function_fb9197e8(L en-US); SetTag("DB_HMI_Ger", 0); SetTag("DB_HMI_Eng/Ger", 1)
   Button "Button_8" at 1687,607 size 160x37; TextOff 'ENGLISH'
      on Click: function_fb9197e8(L en-US); SetTag("DB_HMI_Ger", 0); SetTag("DB_HMI_Eng/Ger", 1)
      Appearance <- "DB_HMI_Eng/Ger"
   Button "Button_9" at 1305,606 size 160x37; TextOff 'DEUTSCH'
      on Click: function_fb9197e8(L de-DE); SetTag("DB_HMI_Ger", 1); SetTag("DB_HMI_Eng/Ger", 0)
      Appearance <- "DB_HMI_Ger"
   GraphicView "Graphic view_24" at 1305,518 size 159x88; Picture "Graphic_126"
   Button "Button_5" at 1305,518 size 159x88; TextOff 'Text'
      on Click: function_fb9197e8(L de-DE); SetTag("DB_HMI_Ger", 1); SetTag("DB_HMI_Eng/Ger", 0)
   TextField "Text field_21" at 1312,143 size 608x40; Text 'REMOTE EMG/STOP/START / FERN-EMG/STOP/START'
   Switch "Switch_2" at 1321,211 size 150x76; TextOn 'EMG'; CaptionText 'Switch'; TextOff 'EMG'
      on SwitchOn: SetTag("DB_RemoteAcces_On/Off", 0)
      Appearance <- "DB_RemoteAcces_EmgStopBtn"
      ProcessValue <- "DB_RemoteAcces_EmgStopBtn"
   Button "Button_3" at 1498,211 size 152x77; TextOff 'Stop'
      on Click: SetTag("DB_RemoteAcces_On/Off", 0)
      Appearance <- "DB_RemoteAcces_On/Off"
      ObjectEnable <- "DB_RemoteAcces_ControlEnable_Stop"
   Button "Button_4" at 1671,212 size 155x76; TextOff 'Start'
      on Click: SetTag("DB_RemoteAcces_On/Off", 1)
      Appearance <- "DB_RemoteAcces_On/Off"
      ObjectEnable <- "DB_RemoteAcces_ControlEnable_Start"
   Switch "Switch_5" at 1325,306 size 255x53; TextOn 'Manual / manuell'; CaptionText 'Switch'; TextOff 'Automat / Automatisch'
      ObjectEnable <- "DB_RemoteAcces_ControlEnable_Man/Auto"
      ProcessValue <- "DB_RemoteAcces_Manual/Auto"
   Switch "Switch_10" at 1593,309 size 233x53; CaptionText 'Switch'; TextOff 'Local / Lokal'; TextOn 'Remote / Fern'; Authorization "Monitor"
      ProcessValue <- "DB_RemoteAcces_Remote"

screen "Statie Incarcare" 1920x1080, template "Template_1"
   GraphicView "Graphic view_4" at 119,0 size 321x185; Picture "background.xwr"
   Rectangle "Rectangle_15" at 191,13 size 169x140
      VerticalMovement <- "DB_general_Poz_Cutie_Bile"
      Visibility <- "DB_Vizibilitati_Platforme/Colete_Platforma_B"
   Rectangle "Rectangle_48" at 191,15 size 169x138
      Visibility <- "DB_HMI_Viz_Platforma_Libera"
      VerticalMovement <- "DB_general_Poz_Cutie_Bile"
   Rectangle "Rectangle_24" at 191,15 size 169x138
      VerticalMovement <- "DB_general_Poz_Cutie_Bile"
      Visibility <- "DB_Vizibilitati_Platforme/Colete_Platforma_A"
   Rectangle "Rectangle_16" at 191,13 size 169x138
      VerticalMovement <- "DB_general_Poz_Cutie_Bile"
      Visibility <- "DB_Vizibilitati_Platforme/Colete_Platforma_C"
   GraphicView "Graphic view_7" at 210,28 size 132x117; Picture "Box"
      VerticalMovement <- "DB_general_Poz_Cutie_Bile"
      Visibility <- "DB_Vizibilitati_Platforme/Colete_Colet_B"
   GraphicView "Graphic view_1" at 210,28 size 132x117; Picture "Box"
      VerticalMovement <- "DB_general_Poz_Cutie_Bile"
      Visibility <- "DB_Vizibilitati_Platforme/Colete_Colet_A"
   GraphicView "Graphic view_6" at 210,28 size 132x117; Picture "Box"
      VerticalMovement <- "DB_general_Poz_Cutie_Bile"
      Visibility <- "DB_Vizibilitati_Platforme/Colete_Colet_C"
   Rectangle "Rectangle_3" at 5,463 size 113x42
      HorizontalMovement <- "DB_general_Piston_Incarcare_B"
   Rectangle "Rectangle_4" at 5,459 size 113x50
      HorizontalMovement <- "DB_general_Piston_Incarcare_B"
   Rectangle "Rectangle_5" at 10,451 size 113x67
      HorizontalMovement <- "DB_general_Piston_Incarcare_B"
   Rectangle "Rectangle_17" at 5,438 size 113x92
      HorizontalMovement <- "DB_general_Piston_Incarcare_B"
   Rectangle "Rectangle_6" at 0,693 size 113x42
      HorizontalMovement <- "DB_general_Piston_Incarcare_C"
   Rectangle "Rectangle_7" at 0,689 size 113x50
      HorizontalMovement <- "DB_general_Piston_Incarcare_C"
   Rectangle "Rectangle_8" at 5,681 size 113x67
      HorizontalMovement <- "DB_general_Piston_Incarcare_C"
   Rectangle "Rectangle_10" at 0,668 size 113x92
      HorizontalMovement <- "DB_general_Piston_Incarcare_C"
   Rectangle "Rectangle_30" at 0,250 size 113x42
      HorizontalMovement <- "DB_general_Piston_Incarcare_A"
   Rectangle "Rectangle_29" at 0,246 size 113x50
      HorizontalMovement <- "DB_general_Piston_Incarcare_A"
   Rectangle "Rectangle_28" at 5,238 size 113x67
      HorizontalMovement <- "DB_general_Piston_Incarcare_A"
   Rectangle "Rectangle_25" at 0,225 size 113x92
      HorizontalMovement <- "DB_general_Piston_Incarcare_A"
   GraphicView "Graphic view_3" at 414,167 size 711x201; Picture "Graphic_30"
   GraphicView "Graphic view_2" at 397,399 size 711x201; Picture "Graphic_30"
   GraphicView "Graphic view_5" at 398,633 size 711x201; Picture "Graphic_30"
   Switch "Switch_1" at 449,34 size 388x100; TextOn 'Transporting / Transport'; CaptionText 'Switch'; TextOff 'Transport'
      on SwitchOn: "VBFunction_4"()
      ProcessValue <- "DB_HMI_Transport"
      Appearance <- "DB_HMI_Transport"
   Rectangle "Rectangle_27" at 102,196 size 38x154
      HorizontalMovement <- "DB_general_Piston_Incarcare_A"
   GraphicView "Graphic view_11" at 9,856 size 162x73; Picture "Graphic_76"
   Rectangle "Rectangle_33" at 77,888 size 45x37
      Appearance <- "DB_HMI_Status_Banda_Bile"
   Rectangle "Rectangle_32" at 107,409 size 38x154
      HorizontalMovement <- "DB_general_Piston_Incarcare_B"
   Rectangle "Rectangle_12" at 102,639 size 38x154
      HorizontalMovement <- "DB_general_Piston_Incarcare_C"
   Rectangle "Rectangle_35" at 27,352 size 107x54
      Appearance <- "DB_Status_Pistoane_Status_Piston_A"
   Rectangle "Rectangle_36" at 29,570 size 107x54
      Appearance <- "DB_Status_Pistoane_Status_Piston_B"
   Rectangle "Rectangle_37" at 31,802 size 107x54
      Appearance <- "DB_Status_Pistoane_Status_Piston_C"
   TextField "Text field_9" at 39,805 size 120x50; Text 'P-C'
   TextField "Text field_11" at 45,574 size 132x50; Text 'P-B'
   TextField "Text field_8" at 39,350 size 120x50; Text 'P-A'
   Button "Button_1" at 848,34 size 239x100; TextOff 'RESET / ZURÜCKSETZEN'
      on Release: SetTag("DB_SIM_BTN_RESET", 0)
      on Press: SetTag("DB_HMI_Viz_Cutie_Scurta", 0); SetTag("LOAD", 0); SetTag("DB_HMI_Ack_Load", 0); SetTag("DB_SIM_BTN_RESET", 1); SetTag("DB_general_Senzor_1_Incarcare", 0); SetTag("DB_general_Senzor_2_Incarcare", 0); SetTag("LOAD", 0); SetTag("DB_HMI_TEST_LOAD", 0); SetTag("DB_HMI_Viz_Cutie_Man/Auto", 0); SetTag("DB_HMI_Viz_Cutie_Banda_1", 0); SetTag("DB_general_Piston_Incarcare_A", 0); SetTag("DB_general_Piston_Incarcare_B", 0); SetTag("DB_general_Piston_Incarcare_C", 0); SetTag("DB_HMI_Cantitate_Loaded_A", 0); SetTag("DB_HMI_Cantitate_Loaded_B", 0); SetTag("DB_HMI_Cantitate_Loaded_C", 0)
      on Click: SetTag("DB_HMI_Total_Weight_A", 0); SetTag("DB_HMI_Total_Weight_B", 0); SetTag("DB_HMI_Total_Weight_C", 0); SetTag("DB_HMI_Cantitate_Loaded_A", 0); SetTag("DB_HMI_Cantitate_Loaded_B", 0); SetTag("DB_HMI_Cantitate_Loaded_C", 0); SetTag("DB_HMI_Total_Weight_A", 0); SetTag("DB_HMI_Total_Weight_B", 0); SetTag("DB_HMI_Total_Weight_C", 0)
   Button "Button_5" at 1120,270 size 178x55; TextOff 'Details Truck A / Details LKW A'
      on Click: SetTag("DB_HMI_Detalii_Truck_A", 1); SetTag("DB_HMI_Detalii_Truck_B", 0); SetTag("DB_HMI_Detalii_Truck_C", 0)
      Appearance <- "DB_HMI_Detalii_Truck_A"
   Button "Button_6" at 1318,270 size 178x55; TextOff 'Details Truck B / Details LKW B'
      on Click: SetTag("DB_HMI_Detalii_Truck_A", 0); SetTag("DB_HMI_Detalii_Truck_B", 1); SetTag("DB_HMI_Detalii_Truck_C", 0)
      Appearance <- "DB_HMI_Detalii_Truck_B"
   Button "Button_7" at 1511,270 size 178x55; TextOff 'Details Truck C / Details LKW C'
      on Click: SetTag("DB_HMI_Detalii_Truck_A", 0); SetTag("DB_HMI_Detalii_Truck_B", 0); SetTag("DB_HMI_Detalii_Truck_C", 1)
      Appearance <- "DB_HMI_Detalii_Truck_C"
   Rectangle "Rectangle_19" at 1128,341 size 550x427
      Visibility <- "DB_HMI_Detalii_Truck_A"
   Rectangle "Rectangle_20" at 1135,347 size 540x76
      Visibility <- "DB_HMI_Detalii_Truck_A"
   TextField "Text field_3" at 1125,369 size 485x40; Text 'Truck A details / Details zum LKW A'
      Visibility <- "DB_HMI_Detalii_Truck_A"
   TextField "Text field_5" at 1079,460 size 397x34; Text 'Available places / Verfügbare Plätze'
      Visibility <- "DB_HMI_Detalii_Truck_A"
   IOField "I/O field_1" at 1521,462 size 96x32; FormatPattern 99
      Visibility <- "DB_HMI_Detalii_Truck_A"
      ProcessValue <- "Locuri_A"
   TextField "Text field_6" at 1087,540 size 389x34; Text 'Loaded packets / Geladene Pakete'
      Visibility <- "DB_HMI_Detalii_Truck_A"
   IOField "I/O field_2" at 1521,538 size 96x32; FormatPattern 99
      ProcessValue <- "DB_HMI_Cantitate_Loaded_A"
      Visibility <- "DB_HMI_Detalii_Truck_A"
   IOField "I/O field_3" at 1247,661 size 124x32; FormatPattern 999; Unit  kg
      ProcessValue <- "DB_HMI_Total_Weight_A"
      Visibility <- "DB_HMI_Detalii_Truck_A"
   IOField "I/O field_4" at 1432,661 size 96x32; FormatPattern 999; Unit  kg
      ProcessValue <- "DB_HMI_MaxLoad_A"
      Visibility <- "DB_HMI_Detalii_Truck_A"
   TextField "Text field_7" at 956,610 size 733x64; Text 'Total weight/ Max weight / Gesamtgewicht/Höchstgewicht'
      Visibility <- "DB_HMI_Detalii_Truck_A"
   TextField "Text field_1" at 192,217 size 645x52; Text 'Truck A / LKW A'
   TextField "Text field_2" at 184,442 size 645x52; Text 'Truck B / LKW B'
   TextField "Text field_14" at 184,678 size 645x52; Text 'Truck C / LKW C'
   TextField "Text field_21" at 1140,25 size 608x40; Text 'REMOTE EMG/STOP/START / FERN-EMG/STOP/START'
   Switch "Switch_2" at 1149,93 size 150x76; TextOn 'EMG'; CaptionText 'Switch'; TextOff 'EMG'
      on SwitchOn: SetTag("DB_RemoteAcces_On/Off", 0)
      Appearance <- "DB_RemoteAcces_EmgStopBtn"
      ProcessValue <- "DB_RemoteAcces_EmgStopBtn"
   Button "Button_3" at 1326,93 size 152x77; TextOff 'Stop'
      on Click: SetTag("DB_RemoteAcces_On/Off", 0)
      Appearance <- "DB_RemoteAcces_On/Off"
      ObjectEnable <- "DB_RemoteAcces_ControlEnable_Stop"
   Button "Button_4" at 1499,94 size 155x76; TextOff 'Start'
      on Click: SetTag("DB_RemoteAcces_On/Off", 1)
      Appearance <- "DB_RemoteAcces_On/Off"
      ObjectEnable <- "DB_RemoteAcces_ControlEnable_Start"
   Switch "Switch_5" at 1153,188 size 255x53; TextOn 'Manual / manuell'; CaptionText 'Switch'; TextOff 'Automat / Automatisch'
      ObjectEnable <- "DB_RemoteAcces_ControlEnable_Man/Auto"
      ProcessValue <- "DB_RemoteAcces_Manual/Auto"
   Switch "Switch_10" at 1421,191 size 233x53; CaptionText 'Switch'; TextOff 'Local / Lokal'; TextOn 'Remote / Fern'; Authorization "Monitor"
      ProcessValue <- "DB_RemoteAcces_Remote"
   Rectangle "Rectangle_9" at 1128,341 size 550x427
      Visibility <- "DB_HMI_Detalii_Truck_B"
   Rectangle "Rectangle_13" at 1135,347 size 540x76
      Visibility <- "DB_HMI_Detalii_Truck_B"
   TextField "Text field_4" at 1125,369 size 485x40; Text 'Truck B details / Details zum LKW B'
      Visibility <- "DB_HMI_Detalii_Truck_B"
   TextField "Text field_10" at 1079,460 size 397x34; Text 'Available places / Verfügbare Plätze'
      Visibility <- "DB_HMI_Detalii_Truck_B"
   IOField "I/O field_5" at 1521,462 size 96x32; FormatPattern 99
      Visibility <- "DB_HMI_Detalii_Truck_B"
      ProcessValue <- "Locuri_B"
   TextField "Text field_12" at 1087,540 size 389x34; Text 'Loaded packets / Geladene Pakete'
      Visibility <- "DB_HMI_Detalii_Truck_B"
   IOField "I/O field_6" at 1521,538 size 96x32; FormatPattern 99
      ProcessValue <- "DB_HMI_Cantitate_Loaded_B"
      Visibility <- "DB_HMI_Detalii_Truck_B"
   TextField "Text field_13" at 956,610 size 733x64; Text 'Total weight/ Max weight / Gesamtgewicht/Höchstgewicht'
      Visibility <- "DB_HMI_Detalii_Truck_B"
   IOField "I/O field_7" at 1275,661 size 96x32; FormatPattern 999; Unit  kg
      ProcessValue <- "DB_HMI_Total_Weight_B"
      Visibility <- "DB_HMI_Detalii_Truck_B"
   IOField "I/O field_8" at 1432,661 size 96x32; FormatPattern 999; Unit  kg
      ProcessValue <- "DB_HMI_MaxLoad_B"
      Visibility <- "DB_HMI_Detalii_Truck_B"
   Rectangle "Rectangle_14" at 1128,341 size 550x426
      Visibility <- "DB_HMI_Detalii_Truck_C"
   Rectangle "Rectangle_18" at 1135,347 size 540x76
      Visibility <- "DB_HMI_Detalii_Truck_C"
   TextField "Text field_16" at 1125,369 size 485x40; Text 'Truck C details / Details zum LKW C'
      Visibility <- "DB_HMI_Detalii_Truck_C"
   TextField "Text field_17" at 1079,460 size 397x34; Text 'Available places / Verfügbare Plätze'
      Visibility <- "DB_HMI_Detalii_Truck_C"
   IOField "I/O field_9" at 1521,462 size 96x32; FormatPattern 99
      Visibility <- "DB_HMI_Detalii_Truck_C"
      ProcessValue <- "Locuri_C"
   TextField "Text field_18" at 1087,540 size 389x34; Text 'Loaded packets / Geladene Pakete'
      Visibility <- "DB_HMI_Detalii_Truck_C"
   IOField "I/O field_10" at 1521,538 size 96x32; FormatPattern 99
      Visibility <- "DB_HMI_Detalii_Truck_C"
      ProcessValue <- "DB_HMI_Cantitate_Loaded_C"
   TextField "Text field_19" at 956,610 size 733x64; Text 'Total weight/ Max weight / Gesamtgewicht/Höchstgewicht'
      Visibility <- "DB_HMI_Detalii_Truck_C"
   IOField "I/O field_11" at 1275,661 size 96x32; FormatPattern 999; Unit  kg
      Visibility <- "DB_HMI_Detalii_Truck_C"
      ProcessValue <- "DB_HMI_Total_Weight_C"
   IOField "I/O field_12" at 1432,661 size 96x32; FormatPattern 999; Unit  kg
      Visibility <- "DB_HMI_Detalii_Truck_C"
      ProcessValue <- "DB_HMI_MaxLoad_C"

screen "Alarme" 1920x1080, template "Template_1"
   AlarmView "Alarm view_2" at 30,42 size 1539x452; ColumnTextAlarmState 'Status'
   AlarmView "Alarm view_1" at 29,503 size 1539x404; ColumnTextAlarmState 'Status'

